// TIA Portal project "Project1Mini Indústria de Engarrafamento Automatizado" (V19)

(* hardware
DEVICE "S7-1200 station_2"  S7-1200 Station
   slot 0: "Rack_0"  S7-1200 Rack  Rack  V1.0
   slot 1: "PLC_1"  CPU 1214C AC/DC/Rly  6ES7 214-1BG40-0XB0  V4.6
DEVICE "HMI_1"  KTP700 Basic PN
   slot 0: "HMI_1"  KTP700 Basic PN  6AV2 123-2GB03-0AX0  17.0.0.0
   slot 1: "HMI_RT_1"  KTP700 Basic PN  6AV2 123-2GB03-0AX0  17.0.0.0
   slot 5: "HMI_1.IE_CP_1"  PROFINET Interface  17.0.0.0
      slot 1: "PROFINET Interface_1"  PROFINET Interface
         slot 1: "Port_1"  Port
*)

// ===== PLC "PLC_1"  CPU 1214C AC/DC/Rly =====

VAR_GLOBAL   // PLC tag table "Default tag table"
   "System_Byte" AT %MB1 : Byte;
   "FirstScan" AT %M1.0 : Bool;
   "DiagStatusUpdate" AT %M1.1 : Bool;
   "AlwaysTRUE" AT %M1.2 : Bool;
   "AlwaysFALSE" AT %M1.3 : Bool;
   "Clock_Byte" AT %MB0 : Byte;
   "Clock_10Hz" AT %M0.0 : Bool;
   "Clock_5Hz" AT %M0.1 : Bool;
   "Clock_2.5Hz" AT %M0.2 : Bool;
   "Clock_2Hz" AT %M0.3 : Bool;
   "Clock_1.25Hz" AT %M0.4 : Bool;
   "Clock_1Hz" AT %M0.5 : Bool;
   "Clock_0.625Hz" AT %M0.6 : Bool;
   "Clock_0.5Hz" AT %M0.7 : Bool;
   "Inciar_Sistema" AT %M2.0 : Bool;
   "Inciar" AT %M2.1 : Bool;
   "Parar" AT %M2.2 : Bool;
   "Ativar_Bomba" AT %M2.3 : Bool;
   "Bomba_Agua" AT %M2.4 : Bool;
   "Nivel_Tanque" AT %MW4 : Int;
   "Acionar_esteira" AT %M2.5 : Bool;
   "esteira" AT %M2.6 : Bool;
   "Movimento_esteira" AT %MW6 : Int;
   "Acionar_Valvula" AT %M2.7 : Bool;
   "Valvula_saida" AT %M3.0 : Bool;
   "Tempo" AT %MD8 : Time;
   "Tempo_saida" AT %MD12 : Time;
   "garrafa_cheia" AT %M3.1 : Bool;
   "Conometro" AT %M3.2 : Bool;
   "garrafas_Lista" AT %MW16 : Int;
END_VAR

// folder: System blocks/Program resources

DATA_BLOCK "IEC_Counter_0_DB"   // DB1
{ S7_Optimized_Access := 'TRUE' }
AUTHOR : Simatic
FAMILY : IEC
NAME : CNTR
VERSION : 1.0
// stored: InstanceOfName IEC_COUNTER
"IEC_COUNTER"
BEGIN
END_DATA_BLOCK

DATA_BLOCK "IEC_Counter_0_DB_1"   // DB2
{ S7_Optimized_Access := 'TRUE' }
AUTHOR : Simatic
FAMILY : IEC
NAME : CNTR
VERSION : 1.0
// stored: InstanceOfName IEC_COUNTER
"IEC_COUNTER"
BEGIN
END_DATA_BLOCK

DATA_BLOCK "IEC_Timer_0_DB"   // DB3
{ S7_Optimized_Access := 'TRUE' }
AUTHOR : Simatic
FAMILY : IEC
NAME : IEC_TMR
VERSION : 1.0
// stored: InstanceOfName IEC_TIMER
"IEC_TIMER"
BEGIN
END_DATA_BLOCK

DATA_BLOCK "IEC_Counter_0_DB_2"   // DB4
{ S7_Optimized_Access := 'TRUE' }
AUTHOR : Simatic
FAMILY : IEC
NAME : CNTR
VERSION : 1.0
// stored: InstanceOfName IEC_COUNTER
"IEC_COUNTER"
BEGIN
END_DATA_BLOCK

// folder: (top level)

ORGANIZATION_BLOCK "Main"   // OB1, LAD, ProgramCycle
TITLE = "Main Program Sweep (Cycle)"
{ S7_Optimized_Access := 'TRUE' }
VERSION : 0.1
   VAR_INPUT
      Initial_Call : Bool;   // Initial call of this OB
      Remanence : Bool;   // =True, if remanent data are available
   END_VAR
BEGIN

REGION Network 1
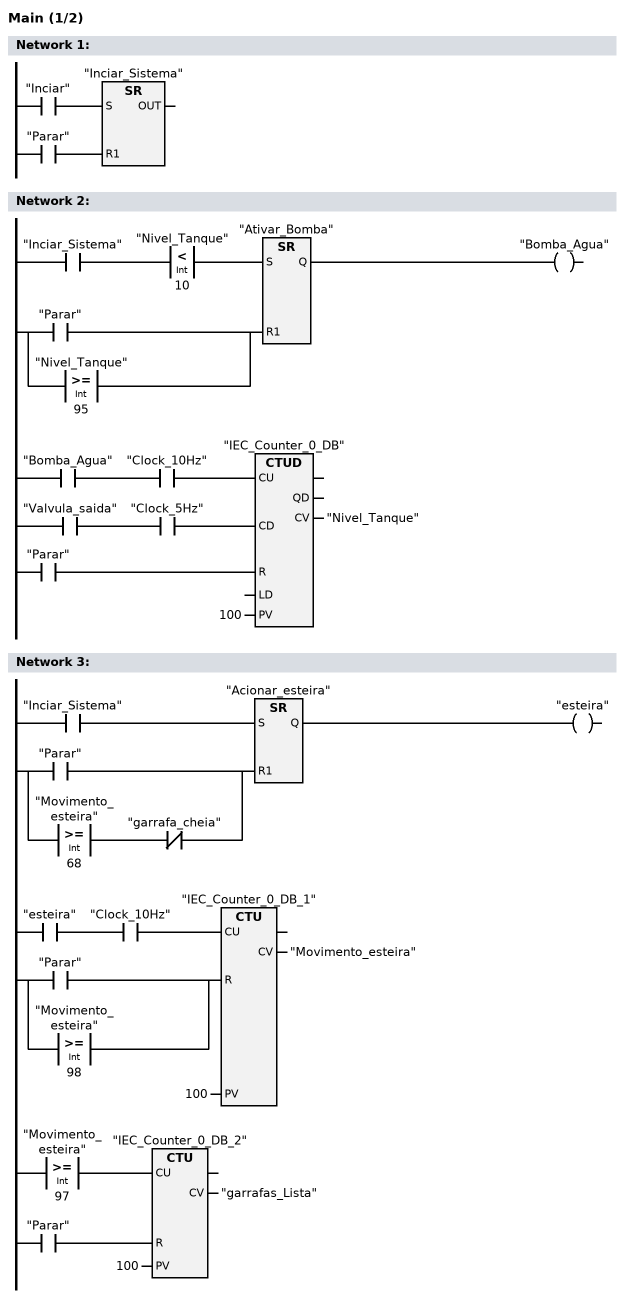
   RUNG wire#powerrail
      Contact( "Inciar" )
      S_SR(operand := "Inciar_Sistema", r1 := wire#w1)
   END_RUNG
   RUNG wire#powerrail
      Contact( "Parar" )
   END_RUNG wire#w1
   // the same network as SCL:
   IF "Inciar" THEN
       "Inciar_Sistema" := TRUE;   // SR flip-flop
   END_IF;
   IF "Parar" THEN "Inciar_Sistema" := FALSE; END_IF;
END_REGION

REGION Network 2
   IF "Inciar_Sistema" AND ("Nivel_Tanque" < 10) THEN
       "Ativar_Bomba" := TRUE;   // SR flip-flop
   END_IF;
   IF "Parar" OR ("Nivel_Tanque" >= 95) THEN "Ativar_Bomba" := FALSE; END_IF;
   "Bomba_Agua" := "Ativar_Bomba";
   "IEC_Counter_0_DB".CTUD(CU := "Bomba_Agua" AND "Clock_10Hz",
                           CD := "Valvula_saida" AND "Clock_5Hz",
                           R := "Parar",
                           PV := 100,
                           CV => "Nivel_Tanque");
END_REGION

REGION Network 3
   IF "Inciar_Sistema" THEN
       "Acionar_esteira" := TRUE;   // SR flip-flop
   END_IF;
   IF "Parar" OR (("Movimento_esteira" >= 68) AND NOT "garrafa_cheia") THEN
       "Acionar_esteira" := FALSE;
   END_IF;
   "esteira" := "Acionar_esteira";
   "IEC_Counter_0_DB_1".CTU(CU := "esteira" AND "Clock_10Hz",
                           R := "Parar" OR ("Movimento_esteira" >= 98),
                           PV := 100,
                           CV => "Movimento_esteira");
   "IEC_Counter_0_DB_2".CTU(CU := "Movimento_esteira" >= 97, R := "Parar", PV := 100, CV => "garrafas_Lista");
END_REGION

REGION Network 4
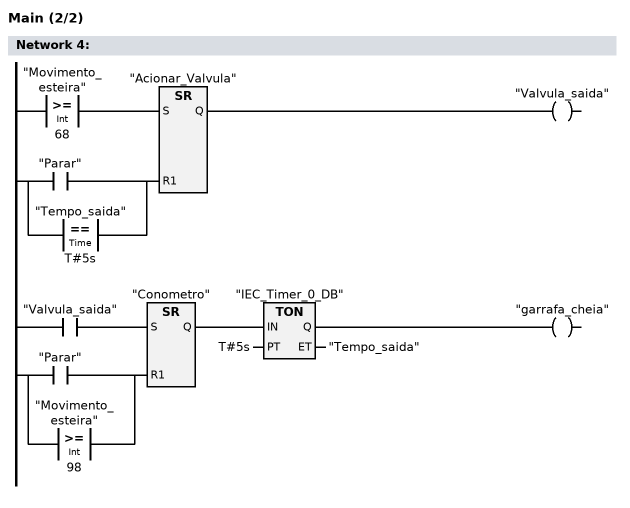
   IF "Movimento_esteira" >= 68 THEN
       "Acionar_Valvula" := TRUE;   // SR flip-flop
   END_IF;
   IF "Parar" OR ("Tempo_saida" = T#5s) THEN "Acionar_Valvula" := FALSE; END_IF;
   "Valvula_saida" := "Acionar_Valvula";
   IF "Valvula_saida" THEN
       "Conometro" := TRUE;   // SR flip-flop
   END_IF;
   IF "Parar" OR ("Movimento_esteira" >= 98) THEN "Conometro" := FALSE; END_IF;
   "IEC_Timer_0_DB".TON(IN := "Conometro", PT := T#5s, ET => "Tempo_saida");
   "garrafa_cheia" := "IEC_Timer_0_DB".Q;
END_REGION
END_ORGANIZATION_BLOCK

(* ===== HMI "HMI_RT_1" =====
system functions are stored by id; their names below are inferred from use
connection "HMI_Connection_1": ETHERNET, SMART_S7_1200_OMS

HMI tags "Default tag table"
   "Tag_ScreenNumber" : UInt, internal
   "Bomba_Agua" : Bool = PLC Bomba_Agua AT %M2.4, 100 ms
   "Nivel_Tanque" : Int = PLC Nivel_Tanque AT %MW4, 100 ms
   "Valvula_saida" : Bool = PLC Valvula_saida AT %M3.0, 100 ms
   "Movimento_esteira" : Int = PLC Movimento_esteira AT %MW6, 100 ms
   "Inciar" : Bool = PLC Inciar AT %M2.1, 100 ms
   "Parar" : Bool = PLC Parar AT %M2.2, 100 ms
   "garrafas_Lista" : Int = PLC garrafas_Lista AT %MW16, 1 s

Template "Template_1" 800x480
   Button "Template_Button" at 714,429 size 71x50; TextOff 'Text'
   Button "Template_Button_1" at 614,429 size 71x50; TextOff 'Text'
   Button "Template_Button_2" at 514,429 size 71x50; TextOff 'Text'
   Button "Template_Button_3" at 414,429 size 71x50; TextOff 'Text'
   Button "Template_Button_4" at 314,429 size 71x50; TextOff 'Text'
   Button "Template_Button_5" at 214,429 size 71x50; TextOff 'Text'
   Button "Alarms" at 114,429 size 71x50; TextOff 'Alarms'; PictureOff "AlarmDisplay_KTP700_Basic_PN_TR"; PictureOn "AlarmDisplay_KTP700_Basic_PN_TR"
      on Release: function_ef3f5d25("Alarm window_Unacknowledged", -1)
   Button "Template_Button_6" at 14,429 size 71x50; TextOff 'Text'
   SymbolicIOField "Symbolic_IO_Field_Screen" at 93,9 size 600x33; TextOff '0'; TextOn '1'; TextList "TextList_ScreenNames"
      ProcessValue <- "Tag_ScreenNumber"
      on Change: ActivateScreenByNumber("Tag_ScreenNumber", 0)
   DateTimeField "HmiScreenItemData" at 695,25 size 105x25
   DateTimeField "HmiScreenItemData_1" at 695,0 size 105x25
   GraphicView "Logo" at 0,0 size 91x51; Picture "Logo of HMI_1"

screen "Root screen" 800x480, template "Template_1"
   on GenerateScreen: SetTag("Tag_ScreenNumber", 1)
   GraphicView "Graphic view_3" at 259,62 size 144x89; Picture "Graphic_7"
   GraphicView "Graphic view_5" at 483,272 size 46x58; Picture "Graphic_9"
   GraphicView "Graphic view_4" at 483,272 size 46x58; Picture "Graphic_8"
      Visibility <- "Valvula_saida"
   GraphicView "Graphic view_9" at 391,42 size 75x75; Picture "Graphic_16"
   GraphicView "Graphic view_2" at 454,37 size 96x245; Picture "Graphic_3"
   GraphicView "Graphic view_1" at 258,62 size 144x89; Picture "Graphic_6"
      Visibility <- "Bomba_Agua"
   Bar "Bar_1" at 466,83 size 74x133; MinimumValue 0; MaximumValue 100
      ProcessValue <- "Nivel_Tanque"
   GraphicView "Graphic view_6" at 2,356 size 798x124; Picture "Graphic_11"
   GraphicView "Graphic view_7" at 125,328 size 52x89; Picture "Graphic_14"
      HorizontalMovement <- "Movimento_esteira"
   Button "Button_2" at 15,142 size 110x52; TextOff 'Parar'
      on Press: SetBit("Parar")
      on Release: ResetBit("Parar")
   Button "Button_1" at 15,71 size 110x52; TextOff 'Inciar'
      on Press: SetBit("Inciar")
      on Release: ResetBit("Inciar")
   Rectangle "Rectangle_3" at 494,350 size 41x58
      Visibility <- "Movimento_esteira"
      HorizontalMovement <- "Movimento_esteira"
   IOField "I/O field_2" at 640,62 size 96x32; FormatPattern 99999
      ProcessValue <- "garrafas_Lista"
*)